// TIA Portal project "FORMING_1500_PLC" (V15) (continued)
REGION Network 33: Control Word Address 12
   RUNG wire#powerrail
      { S7_GenerateENO := "TRUE" } Move(in := 16#047C, out1 => "P_CTW_PROFIBUS_12":P)
   END_RUNG
   // the same network as SCL:
   "P_CTW_PROFIBUS_12":P := 16#047C;
END_REGION

REGION Network 34: Control Word Address 13
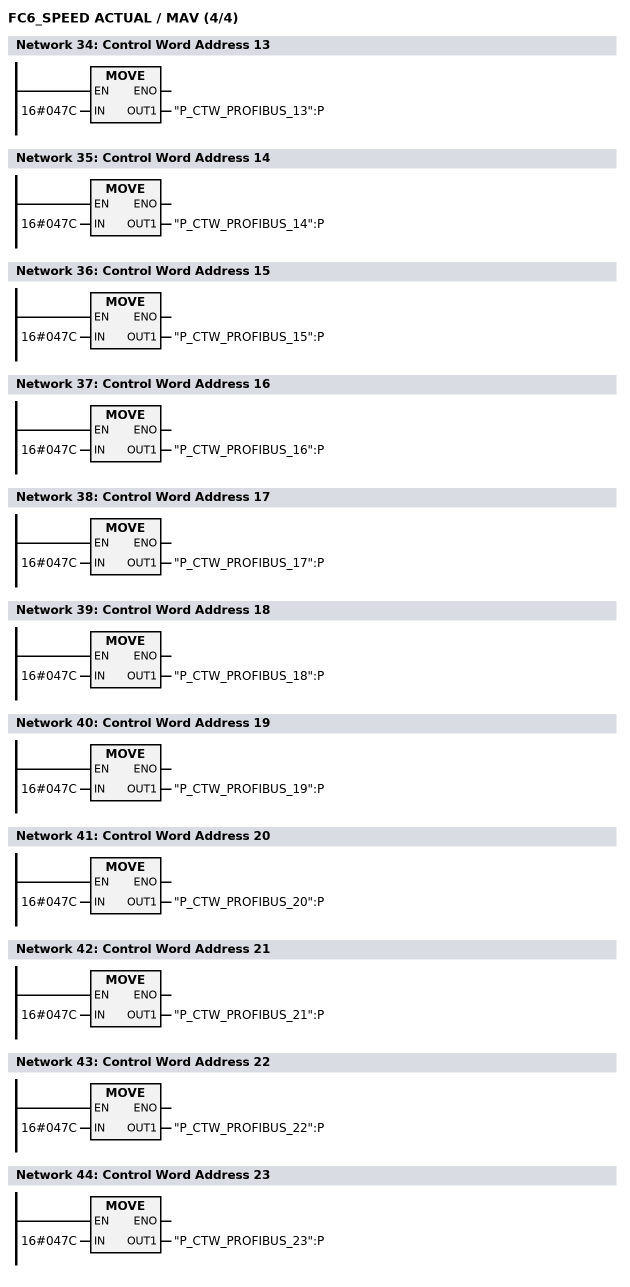
   RUNG wire#powerrail
      { S7_GenerateENO := "TRUE" } Move(in := 16#047C, out1 => "P_CTW_PROFIBUS_13":P)
   END_RUNG
   // the same network as SCL:
   "P_CTW_PROFIBUS_13":P := 16#047C;
END_REGION

REGION Network 35: Control Word Address 14
   RUNG wire#powerrail
      { S7_GenerateENO := "TRUE" } Move(in := 16#047C, out1 => "P_CTW_PROFIBUS_14":P)
   END_RUNG
   // the same network as SCL:
   "P_CTW_PROFIBUS_14":P := 16#047C;
END_REGION

REGION Network 36: Control Word Address 15
   RUNG wire#powerrail
      { S7_GenerateENO := "TRUE" } Move(in := 16#047C, out1 => "P_CTW_PROFIBUS_15":P)
   END_RUNG
   // the same network as SCL:
   "P_CTW_PROFIBUS_15":P := 16#047C;
END_REGION

REGION Network 37: Control Word Address 16
   RUNG wire#powerrail
      { S7_GenerateENO := "TRUE" } Move(in := 16#047C, out1 => "P_CTW_PROFIBUS_16":P)
   END_RUNG
   // the same network as SCL:
   "P_CTW_PROFIBUS_16":P := 16#047C;
END_REGION

REGION Network 38: Control Word Address 17
   RUNG wire#powerrail
      { S7_GenerateENO := "TRUE" } Move(in := 16#047C, out1 => "P_CTW_PROFIBUS_17":P)
   END_RUNG
   // the same network as SCL:
   "P_CTW_PROFIBUS_17":P := 16#047C;
END_REGION

REGION Network 39: Control Word Address 18
   RUNG wire#powerrail
      { S7_GenerateENO := "TRUE" } Move(in := 16#047C, out1 => "P_CTW_PROFIBUS_18":P)
   END_RUNG
   // the same network as SCL:
   "P_CTW_PROFIBUS_18":P := 16#047C;
END_REGION

REGION Network 40: Control Word Address 19
   RUNG wire#powerrail
      { S7_GenerateENO := "TRUE" } Move(in := 16#047C, out1 => "P_CTW_PROFIBUS_19":P)
   END_RUNG
   // the same network as SCL:
   "P_CTW_PROFIBUS_19":P := 16#047C;
END_REGION

REGION Network 41: Control Word Address 20
   RUNG wire#powerrail
      { S7_GenerateENO := "TRUE" } Move(in := 16#047C, out1 => "P_CTW_PROFIBUS_20":P)
   END_RUNG
   // the same network as SCL:
   "P_CTW_PROFIBUS_20":P := 16#047C;
END_REGION

REGION Network 42: Control Word Address 21
   RUNG wire#powerrail
      { S7_GenerateENO := "TRUE" } Move(in := 16#047C, out1 => "P_CTW_PROFIBUS_21":P)
   END_RUNG
   // the same network as SCL:
   "P_CTW_PROFIBUS_21":P := 16#047C;
END_REGION

REGION Network 43: Control Word Address 22
   RUNG wire#powerrail
      { S7_GenerateENO := "TRUE" } Move(in := 16#047C, out1 => "P_CTW_PROFIBUS_22":P)
   END_RUNG
   // the same network as SCL:
   "P_CTW_PROFIBUS_22":P := 16#047C;
END_REGION

REGION Network 44: Control Word Address 23
   RUNG wire#powerrail
      { S7_GenerateENO := "TRUE" } Move(in := 16#047C, out1 => "P_CTW_PROFIBUS_23":P)
   END_RUNG
   // the same network as SCL:
   "P_CTW_PROFIBUS_23":P := 16#047C;
END_REGION
END_FUNCTION

FUNCTION "FC7_INC_DEC_BTN" : Void   // FC7, LAD
TITLE = INCREMENT DECREMENT BUTTN
{ S7_Optimized_Access := 'FALSE' }
VERSION : 0.1
BEGIN

REGION Network 1: METAL DETECT
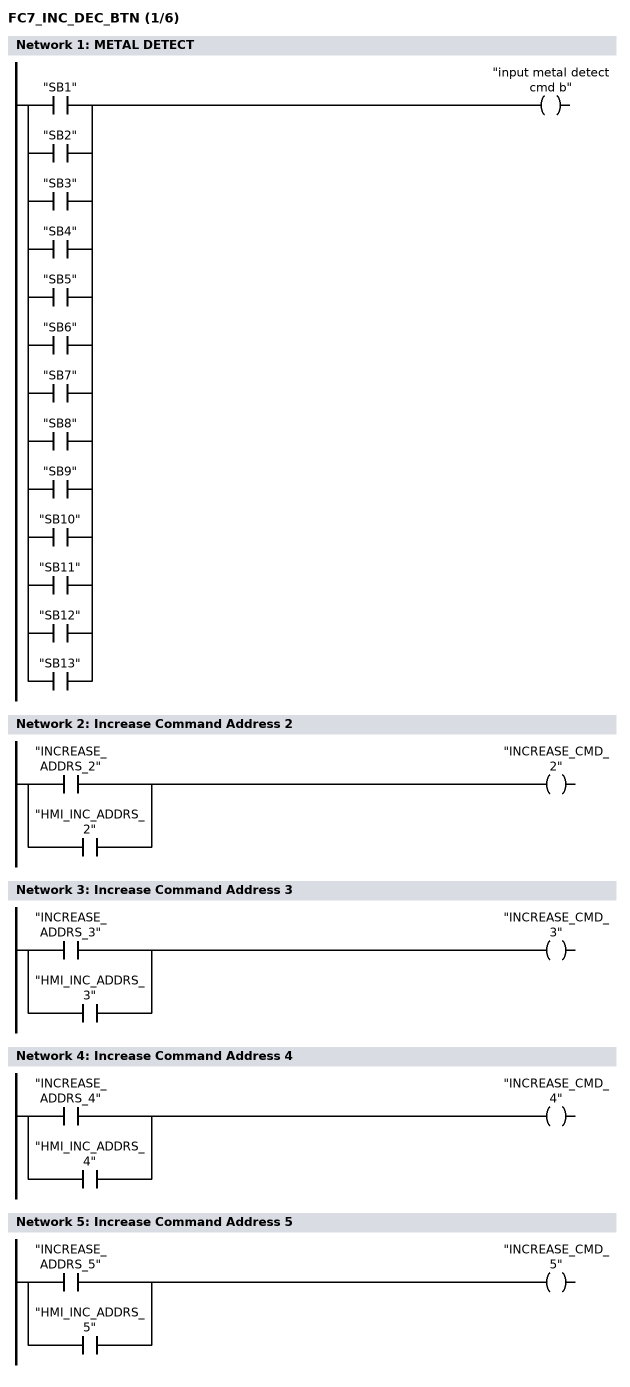
   RUNG wire#powerrail
      Contact( "SB1" )
      wire#w1
      Coil( "input metal detect cmd b" )
   END_RUNG
   RUNG wire#powerrail
      Contact( "SB2" )
   END_RUNG wire#w1
   RUNG wire#powerrail
      Contact( "SB3" )
   END_RUNG wire#w1
   RUNG wire#powerrail
      Contact( "SB4" )
   END_RUNG wire#w1
   RUNG wire#powerrail
      Contact( "SB5" )
   END_RUNG wire#w1
   RUNG wire#powerrail
      Contact( "SB6" )
   END_RUNG wire#w1
   RUNG wire#powerrail
      Contact( "SB7" )
   END_RUNG wire#w1
   RUNG wire#powerrail
      Contact( "SB8" )
   END_RUNG wire#w1
   RUNG wire#powerrail
      Contact( "SB9" )
   END_RUNG wire#w1
   RUNG wire#powerrail
      Contact( "SB10" )
   END_RUNG wire#w1
   RUNG wire#powerrail
      Contact( "SB11" )
   END_RUNG wire#w1
   RUNG wire#powerrail
      Contact( "SB12" )
   END_RUNG wire#w1
   RUNG wire#powerrail
      Contact( "SB13" )
   END_RUNG wire#w1
   // the same network as SCL:
   "input metal detect cmd b" := "SB1" OR "SB2" OR "SB3" OR "SB4" OR "SB5" OR "SB6" OR "SB7" OR "SB8" OR "SB9" OR "SB10" OR "SB11" OR "SB12" OR "SB13";
END_REGION

REGION Network 2: Increase Command Address 2
   RUNG wire#powerrail
      Contact( "INCREASE_ADDRS_2" )
      wire#w1
      Coil( "INCREASE_CMD_2" )
   END_RUNG
   RUNG wire#powerrail
      Contact( "HMI_INC_ADDRS_2" )
   END_RUNG wire#w1
   // the same network as SCL:
   "INCREASE_CMD_2" := "INCREASE_ADDRS_2" OR "HMI_INC_ADDRS_2";
END_REGION

REGION Network 3: Increase Command Address 3
   RUNG wire#powerrail
      Contact( "INCREASE_ADDRS_3" )
      wire#w1
      Coil( "INCREASE_CMD_3" )
   END_RUNG
   RUNG wire#powerrail
      Contact( "HMI_INC_ADDRS_3" )
   END_RUNG wire#w1
   // the same network as SCL:
   "INCREASE_CMD_3" := "INCREASE_ADDRS_3" OR "HMI_INC_ADDRS_3";
END_REGION

REGION Network 4: Increase Command Address 4
   RUNG wire#powerrail
      Contact( "INCREASE_ADDRS_4" )
      wire#w1
      Coil( "INCREASE_CMD_4" )
   END_RUNG
   RUNG wire#powerrail
      Contact( "HMI_INC_ADDRS_4" )
   END_RUNG wire#w1
   // the same network as SCL:
   "INCREASE_CMD_4" := "INCREASE_ADDRS_4" OR "HMI_INC_ADDRS_4";
END_REGION

REGION Network 5: Increase Command Address 5
   RUNG wire#powerrail
      Contact( "INCREASE_ADDRS_5" )
      wire#w1
      Coil( "INCREASE_CMD_5" )
   END_RUNG
   RUNG wire#powerrail
      Contact( "HMI_INC_ADDRS_5" )
   END_RUNG wire#w1
   // the same network as SCL:
   "INCREASE_CMD_5" := "INCREASE_ADDRS_5" OR "HMI_INC_ADDRS_5";
END_REGION

REGION Network 6: Increase Command Address 6
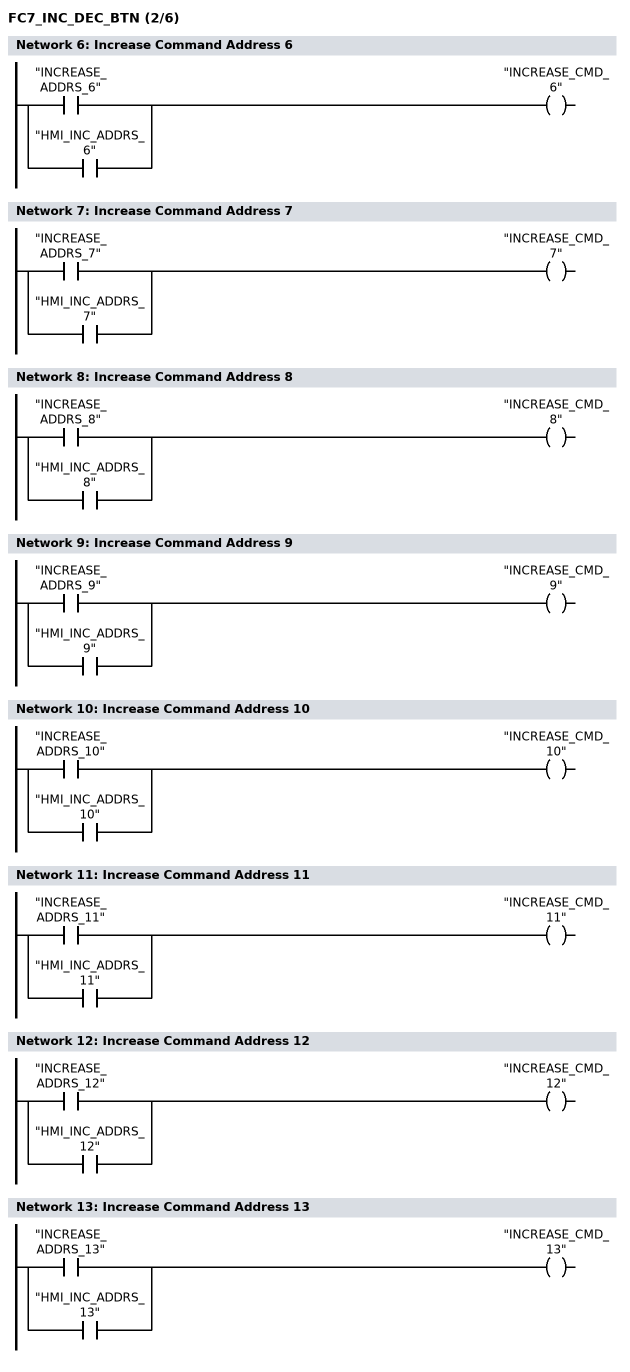
   RUNG wire#powerrail
      Contact( "INCREASE_ADDRS_6" )
      wire#w1
      Coil( "INCREASE_CMD_6" )
   END_RUNG
   RUNG wire#powerrail
      Contact( "HMI_INC_ADDRS_6" )
   END_RUNG wire#w1
   // the same network as SCL:
   "INCREASE_CMD_6" := "INCREASE_ADDRS_6" OR "HMI_INC_ADDRS_6";
END_REGION

REGION Network 7: Increase Command Address 7
   RUNG wire#powerrail
      Contact( "INCREASE_ADDRS_7" )
      wire#w1
      Coil( "INCREASE_CMD_7" )
   END_RUNG
   RUNG wire#powerrail
      Contact( "HMI_INC_ADDRS_7" )
   END_RUNG wire#w1
   // the same network as SCL:
   "INCREASE_CMD_7" := "INCREASE_ADDRS_7" OR "HMI_INC_ADDRS_7";
END_REGION

REGION Network 8: Increase Command Address 8
   RUNG wire#powerrail
      Contact( "INCREASE_ADDRS_8" )
      wire#w1
      Coil( "INCREASE_CMD_8" )
   END_RUNG
   RUNG wire#powerrail
      Contact( "HMI_INC_ADDRS_8" )
   END_RUNG wire#w1
   // the same network as SCL:
   "INCREASE_CMD_8" := "INCREASE_ADDRS_8" OR "HMI_INC_ADDRS_8";
END_REGION

REGION Network 9: Increase Command Address 9
   RUNG wire#powerrail
      Contact( "INCREASE_ADDRS_9" )
      wire#w1
      Coil( "INCREASE_CMD_9" )
   END_RUNG
   RUNG wire#powerrail
      Contact( "HMI_INC_ADDRS_9" )
   END_RUNG wire#w1
   // the same network as SCL:
   "INCREASE_CMD_9" := "INCREASE_ADDRS_9" OR "HMI_INC_ADDRS_9";
END_REGION

REGION Network 10: Increase Command Address 10
   RUNG wire#powerrail
      Contact( "INCREASE_ADDRS_10" )
      wire#w1
      Coil( "INCREASE_CMD_10" )
   END_RUNG
   RUNG wire#powerrail
      Contact( "HMI_INC_ADDRS_10" )
   END_RUNG wire#w1
   // the same network as SCL:
   "INCREASE_CMD_10" := "INCREASE_ADDRS_10" OR "HMI_INC_ADDRS_10";
END_REGION

REGION Network 11: Increase Command Address 11
   RUNG wire#powerrail
      Contact( "INCREASE_ADDRS_11" )
      wire#w1
      Coil( "INCREASE_CMD_11" )
   END_RUNG
   RUNG wire#powerrail
      Contact( "HMI_INC_ADDRS_11" )
   END_RUNG wire#w1
   // the same network as SCL:
   "INCREASE_CMD_11" := "INCREASE_ADDRS_11" OR "HMI_INC_ADDRS_11";
END_REGION

REGION Network 12: Increase Command Address 12
   RUNG wire#powerrail
      Contact( "INCREASE_ADDRS_12" )
      wire#w1
      Coil( "INCREASE_CMD_12" )
   END_RUNG
   RUNG wire#powerrail
      Contact( "HMI_INC_ADDRS_12" )
   END_RUNG wire#w1
   // the same network as SCL:
   "INCREASE_CMD_12" := "INCREASE_ADDRS_12" OR "HMI_INC_ADDRS_12";
END_REGION

REGION Network 13: Increase Command Address 13
   RUNG wire#powerrail
      Contact( "INCREASE_ADDRS_13" )
      wire#w1
      Coil( "INCREASE_CMD_13" )
   END_RUNG
   RUNG wire#powerrail
      Contact( "HMI_INC_ADDRS_13" )
   END_RUNG wire#w1
   // the same network as SCL:
   "INCREASE_CMD_13" := "INCREASE_ADDRS_13" OR "HMI_INC_ADDRS_13";
END_REGION

REGION Network 14: Increase Command Address 14
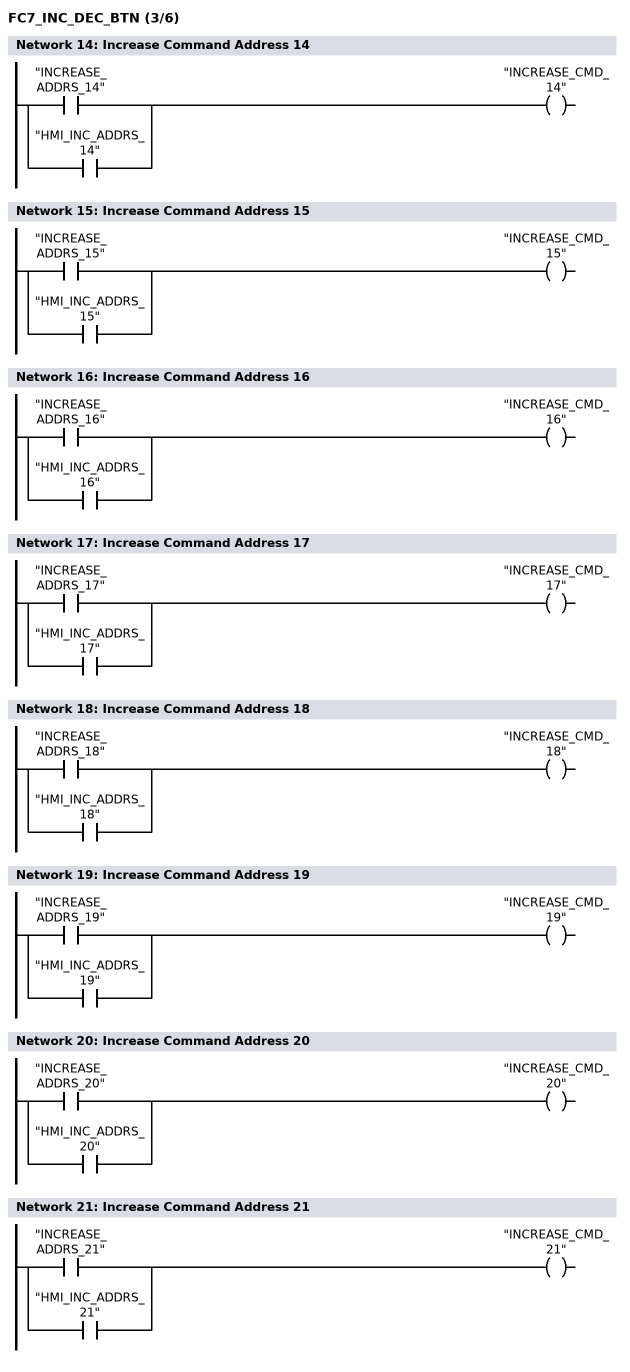
   RUNG wire#powerrail
      Contact( "INCREASE_ADDRS_14" )
      wire#w1
      Coil( "INCREASE_CMD_14" )
   END_RUNG
   RUNG wire#powerrail
      Contact( "HMI_INC_ADDRS_14" )
   END_RUNG wire#w1
   // the same network as SCL:
   "INCREASE_CMD_14" := "INCREASE_ADDRS_14" OR "HMI_INC_ADDRS_14";
END_REGION

REGION Network 15: Increase Command Address 15
   RUNG wire#powerrail
      Contact( "INCREASE_ADDRS_15" )
      wire#w1
      Coil( "INCREASE_CMD_15" )
   END_RUNG
   RUNG wire#powerrail
      Contact( "HMI_INC_ADDRS_15" )
   END_RUNG wire#w1
   // the same network as SCL:
   "INCREASE_CMD_15" := "INCREASE_ADDRS_15" OR "HMI_INC_ADDRS_15";
END_REGION

REGION Network 16: Increase Command Address 16
   RUNG wire#powerrail
      Contact( "INCREASE_ADDRS_16" )
      wire#w1
      Coil( "INCREASE_CMD_16" )
   END_RUNG
   RUNG wire#powerrail
      Contact( "HMI_INC_ADDRS_16" )
   END_RUNG wire#w1
   // the same network as SCL:
   "INCREASE_CMD_16" := "INCREASE_ADDRS_16" OR "HMI_INC_ADDRS_16";
END_REGION

REGION Network 17: Increase Command Address 17
   RUNG wire#powerrail
      Contact( "INCREASE_ADDRS_17" )
      wire#w1
      Coil( "INCREASE_CMD_17" )
   END_RUNG
   RUNG wire#powerrail
      Contact( "HMI_INC_ADDRS_17" )
   END_RUNG wire#w1
   // the same network as SCL:
   "INCREASE_CMD_17" := "INCREASE_ADDRS_17" OR "HMI_INC_ADDRS_17";
END_REGION

REGION Network 18: Increase Command Address 18
   RUNG wire#powerrail
      Contact( "INCREASE_ADDRS_18" )
      wire#w1
      Coil( "INCREASE_CMD_18" )
   END_RUNG
   RUNG wire#powerrail
      Contact( "HMI_INC_ADDRS_18" )
   END_RUNG wire#w1
   // the same network as SCL:
   "INCREASE_CMD_18" := "INCREASE_ADDRS_18" OR "HMI_INC_ADDRS_18";
END_REGION

REGION Network 19: Increase Command Address 19
   RUNG wire#powerrail
      Contact( "INCREASE_ADDRS_19" )
      wire#w1
      Coil( "INCREASE_CMD_19" )
   END_RUNG
   RUNG wire#powerrail
      Contact( "HMI_INC_ADDRS_19" )
   END_RUNG wire#w1
   // the same network as SCL:
   "INCREASE_CMD_19" := "INCREASE_ADDRS_19" OR "HMI_INC_ADDRS_19";
END_REGION

REGION Network 20: Increase Command Address 20
   RUNG wire#powerrail
      Contact( "INCREASE_ADDRS_20" )
      wire#w1
      Coil( "INCREASE_CMD_20" )
   END_RUNG
   RUNG wire#powerrail
      Contact( "HMI_INC_ADDRS_20" )
   END_RUNG wire#w1
   // the same network as SCL:
   "INCREASE_CMD_20" := "INCREASE_ADDRS_20" OR "HMI_INC_ADDRS_20";
END_REGION

REGION Network 21: Increase Command Address 21
   RUNG wire#powerrail
      Contact( "INCREASE_ADDRS_21" )
      wire#w1
      Coil( "INCREASE_CMD_21" )
   END_RUNG
   RUNG wire#powerrail
      Contact( "HMI_INC_ADDRS_21" )
   END_RUNG wire#w1
   // the same network as SCL:
   "INCREASE_CMD_21" := "INCREASE_ADDRS_21" OR "HMI_INC_ADDRS_21";
END_REGION

REGION Network 22: Increase Command Address 22
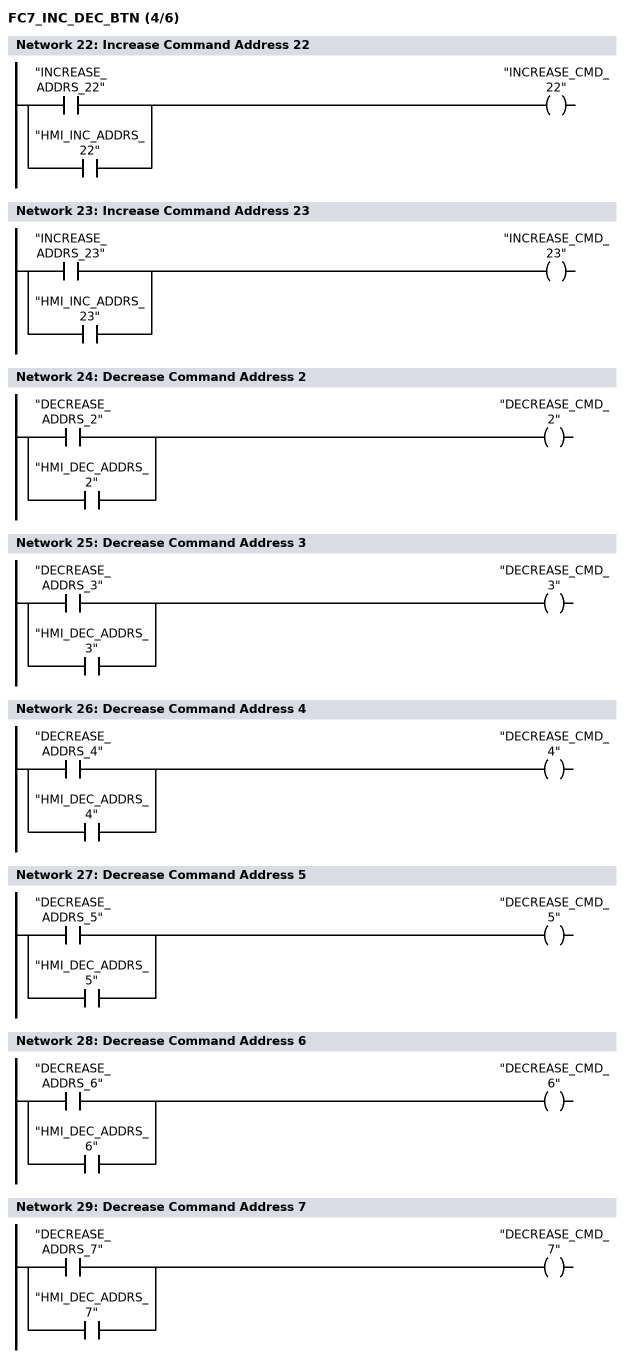
   RUNG wire#powerrail
      Contact( "INCREASE_ADDRS_22" )
      wire#w1
      Coil( "INCREASE_CMD_22" )
   END_RUNG
   RUNG wire#powerrail
      Contact( "HMI_INC_ADDRS_22" )
   END_RUNG wire#w1
   // the same network as SCL:
   "INCREASE_CMD_22" := "INCREASE_ADDRS_22" OR "HMI_INC_ADDRS_22";
END_REGION

REGION Network 23: Increase Command Address 23
   RUNG wire#powerrail
      Contact( "INCREASE_ADDRS_23" )
      wire#w1
      Coil( "INCREASE_CMD_23" )
   END_RUNG
   RUNG wire#powerrail
      Contact( "HMI_INC_ADDRS_23" )
   END_RUNG wire#w1
   // the same network as SCL:
   "INCREASE_CMD_23" := "INCREASE_ADDRS_23" OR "HMI_INC_ADDRS_23";
END_REGION

REGION Network 24: Decrease Command Address 2
   RUNG wire#powerrail
      Contact( "DECREASE_ADDRS_2" )
      wire#w1
      Coil( "DECREASE_CMD_2" )
   END_RUNG
   RUNG wire#powerrail
      Contact( "HMI_DEC_ADDRS_2" )
   END_RUNG wire#w1
   // the same network as SCL:
   "DECREASE_CMD_2" := "DECREASE_ADDRS_2" OR "HMI_DEC_ADDRS_2";
END_REGION

REGION Network 25: Decrease Command Address 3
   RUNG wire#powerrail
      Contact( "DECREASE_ADDRS_3" )
      wire#w1
      Coil( "DECREASE_CMD_3" )
   END_RUNG
   RUNG wire#powerrail
      Contact( "HMI_DEC_ADDRS_3" )
   END_RUNG wire#w1
   // the same network as SCL:
   "DECREASE_CMD_3" := "DECREASE_ADDRS_3" OR "HMI_DEC_ADDRS_3";
END_REGION

REGION Network 26: Decrease Command Address 4
   RUNG wire#powerrail
      Contact( "DECREASE_ADDRS_4" )
      wire#w1
      Coil( "DECREASE_CMD_4" )
   END_RUNG
   RUNG wire#powerrail
      Contact( "HMI_DEC_ADDRS_4" )
   END_RUNG wire#w1
   // the same network as SCL:
   "DECREASE_CMD_4" := "DECREASE_ADDRS_4" OR "HMI_DEC_ADDRS_4";
END_REGION

REGION Network 27: Decrease Command Address 5
   RUNG wire#powerrail
      Contact( "DECREASE_ADDRS_5" )
      wire#w1
      Coil( "DECREASE_CMD_5" )
   END_RUNG
   RUNG wire#powerrail
      Contact( "HMI_DEC_ADDRS_5" )
   END_RUNG wire#w1
   // the same network as SCL:
   "DECREASE_CMD_5" := "DECREASE_ADDRS_5" OR "HMI_DEC_ADDRS_5";
END_REGION

REGION Network 28: Decrease Command Address 6
   RUNG wire#powerrail
      Contact( "DECREASE_ADDRS_6" )
      wire#w1
      Coil( "DECREASE_CMD_6" )
   END_RUNG
   RUNG wire#powerrail
      Contact( "HMI_DEC_ADDRS_6" )
   END_RUNG wire#w1
   // the same network as SCL:
   "DECREASE_CMD_6" := "DECREASE_ADDRS_6" OR "HMI_DEC_ADDRS_6";
END_REGION

REGION Network 29: Decrease Command Address 7
   RUNG wire#powerrail
      Contact( "DECREASE_ADDRS_7" )
      wire#w1
      Coil( "DECREASE_CMD_7" )
   END_RUNG
   RUNG wire#powerrail
      Contact( "HMI_DEC_ADDRS_7" )
   END_RUNG wire#w1
   // the same network as SCL:
   "DECREASE_CMD_7" := "DECREASE_ADDRS_7" OR "HMI_DEC_ADDRS_7";
END_REGION

REGION Network 30: Decrease Command Address 8
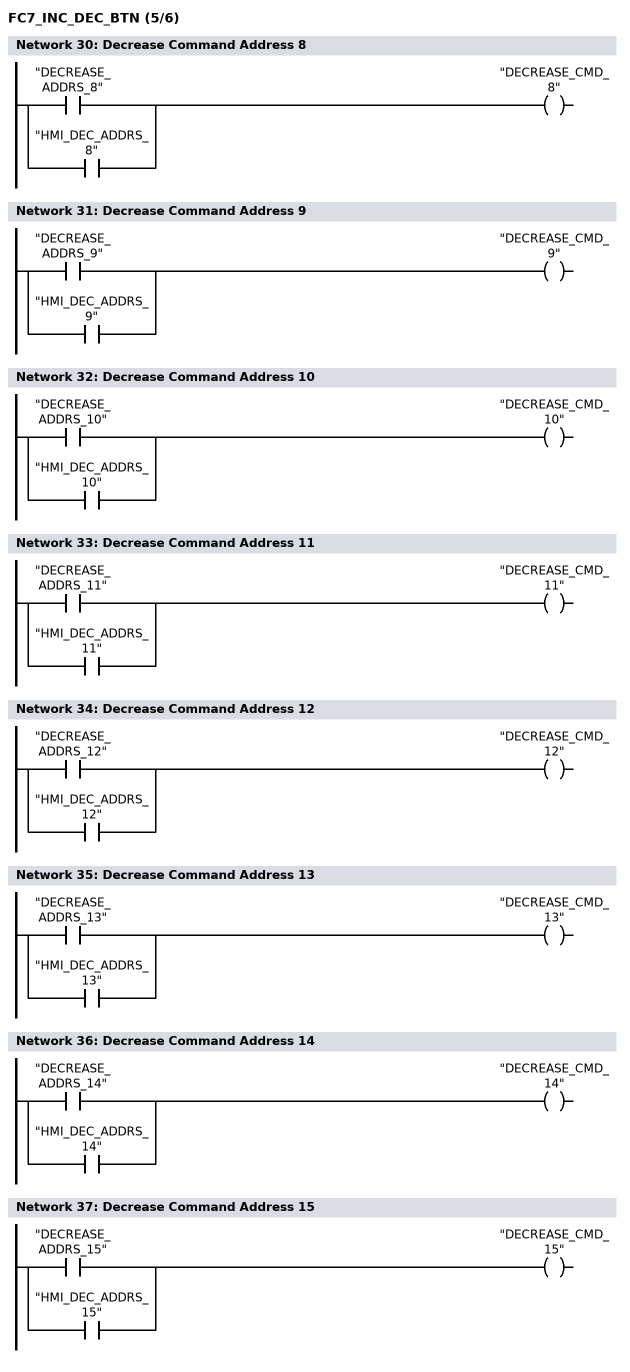
   RUNG wire#powerrail
      Contact( "DECREASE_ADDRS_8" )
      wire#w1
      Coil( "DECREASE_CMD_8" )
   END_RUNG
   RUNG wire#powerrail
      Contact( "HMI_DEC_ADDRS_8" )
   END_RUNG wire#w1
   // the same network as SCL:
   "DECREASE_CMD_8" := "DECREASE_ADDRS_8" OR "HMI_DEC_ADDRS_8";
END_REGION

REGION Network 31: Decrease Command Address 9
   RUNG wire#powerrail
      Contact( "DECREASE_ADDRS_9" )
      wire#w1
      Coil( "DECREASE_CMD_9" )
   END_RUNG
   RUNG wire#powerrail
      Contact( "HMI_DEC_ADDRS_9" )
   END_RUNG wire#w1
   // the same network as SCL:
   "DECREASE_CMD_9" := "DECREASE_ADDRS_9" OR "HMI_DEC_ADDRS_9";
END_REGION

REGION Network 32: Decrease Command Address 10
   RUNG wire#powerrail
      Contact( "DECREASE_ADDRS_10" )
      wire#w1
      Coil( "DECREASE_CMD_10" )
   END_RUNG
   RUNG wire#powerrail
      Contact( "HMI_DEC_ADDRS_10" )
   END_RUNG wire#w1
   // the same network as SCL:
   "DECREASE_CMD_10" := "DECREASE_ADDRS_10" OR "HMI_DEC_ADDRS_10";
END_REGION

REGION Network 33: Decrease Command Address 11
   RUNG wire#powerrail
      Contact( "DECREASE_ADDRS_11" )
      wire#w1
      Coil( "DECREASE_CMD_11" )
   END_RUNG
   RUNG wire#powerrail
      Contact( "HMI_DEC_ADDRS_11" )
   END_RUNG wire#w1
   // the same network as SCL:
   "DECREASE_CMD_11" := "DECREASE_ADDRS_11" OR "HMI_DEC_ADDRS_11";
END_REGION

REGION Network 34: Decrease Command Address 12
   RUNG wire#powerrail
      Contact( "DECREASE_ADDRS_12" )
      wire#w1
      Coil( "DECREASE_CMD_12" )
   END_RUNG
   RUNG wire#powerrail
      Contact( "HMI_DEC_ADDRS_12" )
   END_RUNG wire#w1
   // the same network as SCL:
   "DECREASE_CMD_12" := "DECREASE_ADDRS_12" OR "HMI_DEC_ADDRS_12";
END_REGION

REGION Network 35: Decrease Command Address 13
   RUNG wire#powerrail
      Contact( "DECREASE_ADDRS_13" )
      wire#w1
      Coil( "DECREASE_CMD_13" )
   END_RUNG
   RUNG wire#powerrail
      Contact( "HMI_DEC_ADDRS_13" )
   END_RUNG wire#w1
   // the same network as SCL:
   "DECREASE_CMD_13" := "DECREASE_ADDRS_13" OR "HMI_DEC_ADDRS_13";
END_REGION

REGION Network 36: Decrease Command Address 14
   RUNG wire#powerrail
      Contact( "DECREASE_ADDRS_14" )
      wire#w1
      Coil( "DECREASE_CMD_14" )
   END_RUNG
   RUNG wire#powerrail
      Contact( "HMI_DEC_ADDRS_14" )
   END_RUNG wire#w1
   // the same network as SCL:
   "DECREASE_CMD_14" := "DECREASE_ADDRS_14" OR "HMI_DEC_ADDRS_14";
END_REGION

REGION Network 37: Decrease Command Address 15
   RUNG wire#powerrail
      Contact( "DECREASE_ADDRS_15" )
      wire#w1
      Coil( "DECREASE_CMD_15" )
   END_RUNG
   RUNG wire#powerrail
      Contact( "HMI_DEC_ADDRS_15" )
   END_RUNG wire#w1
   // the same network as SCL:
   "DECREASE_CMD_15" := "DECREASE_ADDRS_15" OR "HMI_DEC_ADDRS_15";
END_REGION

REGION Network 38: Decrease Command Address 16
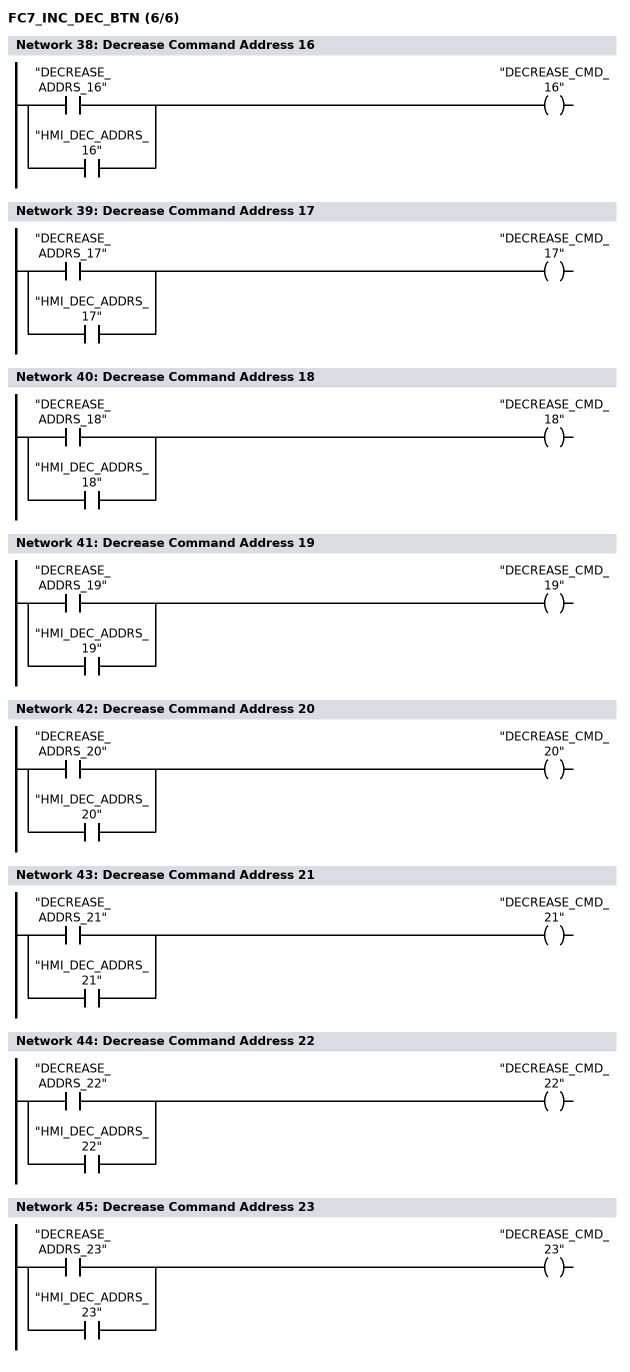
   RUNG wire#powerrail
      Contact( "DECREASE_ADDRS_16" )
      wire#w1
      Coil( "DECREASE_CMD_16" )
   END_RUNG
   RUNG wire#powerrail
      Contact( "HMI_DEC_ADDRS_16" )
   END_RUNG wire#w1
   // the same network as SCL:
   "DECREASE_CMD_16" := "DECREASE_ADDRS_16" OR "HMI_DEC_ADDRS_16";
END_REGION

REGION Network 39: Decrease Command Address 17
   RUNG wire#powerrail
      Contact( "DECREASE_ADDRS_17" )
      wire#w1
      Coil( "DECREASE_CMD_17" )
   END_RUNG
   RUNG wire#powerrail
      Contact( "HMI_DEC_ADDRS_17" )
   END_RUNG wire#w1
   // the same network as SCL:
   "DECREASE_CMD_17" := "DECREASE_ADDRS_17" OR "HMI_DEC_ADDRS_17";
END_REGION

REGION Network 40: Decrease Command Address 18
   RUNG wire#powerrail
      Contact( "DECREASE_ADDRS_18" )
      wire#w1
      Coil( "DECREASE_CMD_18" )
   END_RUNG
   RUNG wire#powerrail
      Contact( "HMI_DEC_ADDRS_18" )
   END_RUNG wire#w1
   // the same network as SCL:
   "DECREASE_CMD_18" := "DECREASE_ADDRS_18" OR "HMI_DEC_ADDRS_18";
END_REGION

REGION Network 41: Decrease Command Address 19
   RUNG wire#powerrail
      Contact( "DECREASE_ADDRS_19" )
      wire#w1
      Coil( "DECREASE_CMD_19" )
   END_RUNG
   RUNG wire#powerrail
      Contact( "HMI_DEC_ADDRS_19" )
   END_RUNG wire#w1
   // the same network as SCL:
   "DECREASE_CMD_19" := "DECREASE_ADDRS_19" OR "HMI_DEC_ADDRS_19";
END_REGION

REGION Network 42: Decrease Command Address 20
   RUNG wire#powerrail
      Contact( "DECREASE_ADDRS_20" )
      wire#w1
      Coil( "DECREASE_CMD_20" )
   END_RUNG
   RUNG wire#powerrail
      Contact( "HMI_DEC_ADDRS_20" )
   END_RUNG wire#w1
   // the same network as SCL:
   "DECREASE_CMD_20" := "DECREASE_ADDRS_20" OR "HMI_DEC_ADDRS_20";
END_REGION

REGION Network 43: Decrease Command Address 21
   RUNG wire#powerrail
      Contact( "DECREASE_ADDRS_21" )
      wire#w1
      Coil( "DECREASE_CMD_21" )
   END_RUNG
   RUNG wire#powerrail
      Contact( "HMI_DEC_ADDRS_21" )
   END_RUNG wire#w1
   // the same network as SCL:
   "DECREASE_CMD_21" := "DECREASE_ADDRS_21" OR "HMI_DEC_ADDRS_21";
END_REGION

REGION Network 44: Decrease Command Address 22
   RUNG wire#powerrail
      Contact( "DECREASE_ADDRS_22" )
      wire#w1
      Coil( "DECREASE_CMD_22" )
   END_RUNG
   RUNG wire#powerrail
      Contact( "HMI_DEC_ADDRS_22" )
   END_RUNG wire#w1
   // the same network as SCL:
   "DECREASE_CMD_22" := "DECREASE_ADDRS_22" OR "HMI_DEC_ADDRS_22";
END_REGION

REGION Network 45: Decrease Command Address 23
   RUNG wire#powerrail
      Contact( "DECREASE_ADDRS_23" )
      wire#w1
      Coil( "DECREASE_CMD_23" )
   END_RUNG
   RUNG wire#powerrail
      Contact( "HMI_DEC_ADDRS_23" )
   END_RUNG wire#w1
   // the same network as SCL:
   "DECREASE_CMD_23" := "DECREASE_ADDRS_23" OR "HMI_DEC_ADDRS_23";
END_REGION
END_FUNCTION

FUNCTION "FC8_SCALLING MAV" : Void   // FC8, LAD
TITLE = SCALLING SPEED ACTUAL FROM INVERTER
{ S7_Optimized_Access := 'FALSE' }
VERSION : 0.1
BEGIN

REGION Network 1: ADDRESS 2
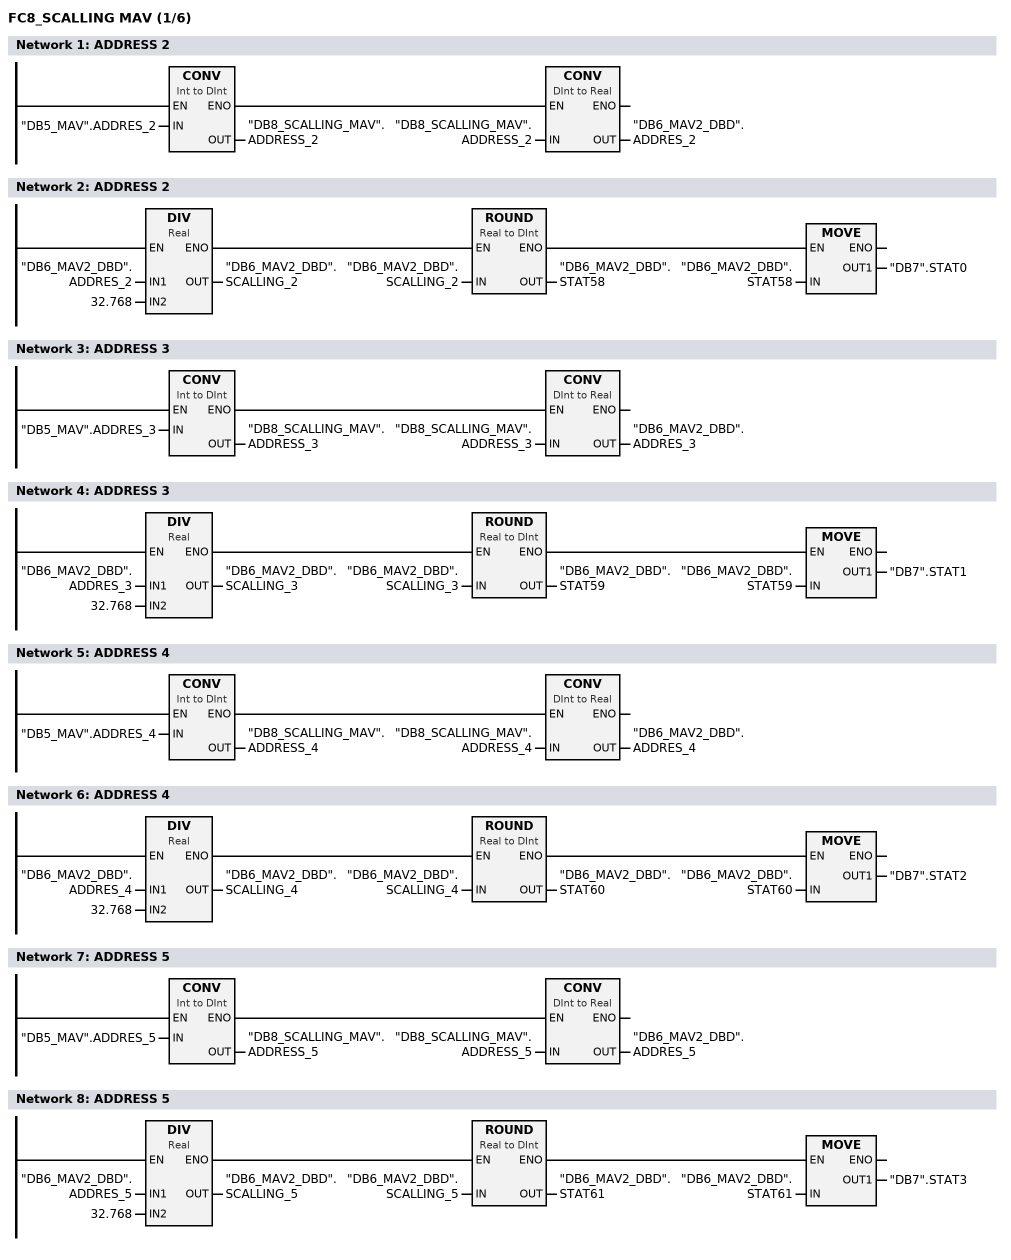
   RUNG wire#powerrail
      { S7_Templates := "[SrcType := Int, DestType := DInt]"; S7_GenerateENO := "TRUE" } Convert(in := "DB5_MAV".ADDRES_2, out => "DB8_SCALLING_MAV".ADDRESS_2)
      { S7_Templates := "[SrcType := DInt, DestType := Real]"; S7_GenerateENO := "TRUE" } Convert(in := "DB8_SCALLING_MAV".ADDRESS_2, out => "DB6_MAV2_DBD".ADDRES_2)
   END_RUNG
   // the same network as SCL:
   // ENO of a box is taken as its EN; it also drops when the box reports an error
   "DB8_SCALLING_MAV".ADDRESS_2 := INT_TO_DINT("DB5_MAV".ADDRES_2);
   "DB6_MAV2_DBD".ADDRES_2 := DINT_TO_REAL("DB8_SCALLING_MAV".ADDRESS_2);
END_REGION

